(* Logix 5000 project; controller POA Emulate 5570 rev 30.12; software revision 30.00 *)

TASK MainTask (periodic, rate 10000 ms, priority 1, watchdog 10000 ms) : MainProgram

MODULES
   Local : Emulate 5570 (ICP 2, rev 30.12)
END_MODULES

VAR_GLOBAL   (* controller tags *)
   _SEC_P : BOOL;
   done : DINT;
   R_TRIG : FBD_ONESHOT;
   temp_var : DINT;
   test_array : DINT[20] := ([0] := 1, [1] := 2, [2] := 3, [3] := 4, [4] := 5, [5] := 6, [6] := 7, [7] := 8, [8] := 9, [9] := 10, [10] := 11, [11] := 12, [12] := 13, [13] := 14, [14] := 15, [15] := 16, [16] := 17, [17] := 18, [18] := 19, [19] := 20);
   TON : FBD_TIMER;
END_VAR

PROGRAM MainProgram   (* main routine MainRoutine *)
VAR
   Chaskey_128_i : DINT;
   Chaskey_a : DINT; {access None}
   Chaskey_BNum : DINT; {access None}
   Chaskey_i : DINT; {access None}
   Chaskey_IndexDiv : DINT;
   Chaskey_IndexMod : DINT;
   Chaskey_input_pi : DINT[4]; {access None}
   Chaskey_j : DINT; {access None}
   Chaskey_key : DINT[4]; {access None}
   Chaskey_L : DINT[4]; {access None}
   Chaskey_LastBlk : DINT[4];
   Chaskey_lb : DINT[16];
   Chaskey_Message : DINT[256]; {access None}
   Chaskey_mlen : DINT;
   Chaskey_MsgBitLen : DINT;
   Chaskey_MsgBlk : DINT[16];
   Chaskey_MsgBlkLen : DINT;
   Chaskey_per_i : DINT; {access None}
   Chaskey_round : DINT;
   Chaskey_shift_input : DINT; {access None}
   Chaskey_shift_result : DINT; {access None}
   Chaskey_subkey1_i : DINT; {access None}
   Chaskey_subkey2_i : DINT; {access None}
   Chaskey_subkey_1 : DINT[8];
   Chaskey_subkey_2 : DINT[8]; {access None}
   Chaskey_tag : DINT[4]; {access None}
   Chaskey_Temp : DINT; {access None}
   Chaskey_z : DINT;
   Date_time : DINT[7]; {access None}
        [0]   // Year
        [1]   // Month
        [2]   // Day
        [3]   // Hour
        [4]   // Minute
        [5]   // Second
        [6]   // Microsecond
   OWF_Add_c : DINT;
   OWF_i : DINT;
   OWF_Input : DINT[17];
   OWF_InputLen : DINT;
   OWF_InputMaxInd : DINT;
   OWF_Result : DINT[17];
   POA_Chain_NM : DINT; {access None}
   POA_CK_RefillNM : DINT; {access None}
   POA_CKP : DINT[17]; {access None}
   POA_CKP_Ctx : DINT[9,16]; {access None}
   POA_CKP_Indx : DINT[9]; {access None}
   POA_i : DINT;
   POA_Ins_NM : DINT; {access None}
   POA_is_Bootstrap : BOOL; {access None}
   POA_j : DINT;
   POA_k : DINT; {access None}
   POA_lr : DINT;
   POA_m : DINT;
   POA_Microsecond1 : DINT; {access None}
   POA_Microsecond2 : DINT; {access None}
   POA_MicrosecondABS : DINT;
   POA_OTS : SINT[256,256];
   POA_Pf : DINT[17]; {access None}
   POA_Pf_Indx : DINT; {access None}
   PoA_Pf_Interval : DINT;
   POA_Qu_head : DINT; {access None}
   POA_Qu_tail : DINT; {access None}
   POA_SC_DeltaS : DINT;
   POA_SC_Interval : DINT;
   POA_Second1 : DINT; {access None}
   POA_Second2 : DINT; {access None}
   POA_SecondABS : DINT;
   POA_SIG_i : DINT;
   POA_tag : DINT[4]; {access None}
   POA_Vrf_Points : DINT[260,17];
   PRG_Counter : DINT[2];
   PRG_i : DINT;
   PRG_j : DINT;
   PRG_Res_Len : DINT;
   PRG_Result : DINT[128];
   SCAN_CYCLE_TIME : DINT; {access None}
   UOWHF_Add_c : DINT;
   UOWHF_i : DINT;
   UOWHF_InputLen : DINT;
   UOWHF_InputMaxInd : DINT := 7;
   UOWHF_Msg : DINT[17];
   UOWHF_OutputMaxInd : DINT;
   UOWHF_Result : DINT[17];
   UOWHF_Vary_BlkNum : DINT;
   UOWHF_Vary_i : DINT := 256;
   UOWHF_Vary_j : DINT;
   UOWHF_Vary_Message : DINT[3000] := ([0] := 1, [1] := 1, [2] := 1, [3] := 1, [4] := 1, [5] := 1, [6] := 1, [7] := 1, [8] := 1, [9] := 1, [10] := 1, [11] := 1, [12] := 1, [13] := 1, [14] := 1, [15] := 1, [16] := 1, [17] := 1, [18] := 1, [19] := 1, [20] := 1, [21] := 1, [22] := 1, [23] := 1, [24] := 1, [25] := 1, [26] := 1, [27] := 1, [28] := 1, [29] := 1, [30] := 1, [31] := 1, [32] := 1, [33] := 1, [34] := 1, [35] := 1, [36] := 1, [37] := 1, [38] := 1, [39] := 1, [40] := 1, [41] := 1, [42] := 1, [43] := 1, [44] := 1, [45] := 1, [46] := 1, [47] := 1, [48] := 1, [49] := 1, [50] := 1, [51] := 1, [52] := 1, [53] := 1, [54] := 1, [55] := 1, [56] := 1, [57] := 1, [58] := 1, [59] := 1,
        [60] := 1, [61] := 1, [62] := 1, [63] := 1, [64] := 1, [65] := 1, [66] := 1, [67] := 1, [68] := 1, [69] := 1, [70] := 1, [71] := 1, [72] := 1, [73] := 1, [74] := 1, [75] := 1, [76] := 1, [77] := 1, [78] := 1, [79] := 1, [80] := 1, [81] := 1, [82] := 1, [83] := 1, [84] := 1, [85] := 1, [86] := 1, [87] := 1, [88] := 1, [89] := 1, [90] := 1, [91] := 1, [92] := 1, [93] := 1, [94] := 1, [95] := 1, [96] := 1, [97] := 1, [98] := 1, [99] := 1, [100] := 1, [101] := 1, [102] := 1, [103] := 1, [104] := 1, [105] := 1, [106] := 1, [107] := 1, [108] := 1, [109] := 1, [110] := 1, [111] := 1, [112] := 1, [113] := 1, [114] := 1, [115] := 1, [116] := 1, [117] := 1, [118] := 1, [119] := 1,
        [120] := 1, [121] := 1, [122] := 1, [123] := 1, [124] := 1, [125] := 1, [126] := 1, [127] := 1, [128] := 1, [129] := 1, [130] := 1, [131] := 1, [132] := 1, [133] := 1, [134] := 1, [135] := 1, [136] := 1, [137] := 1, [138] := 1, [139] := 1, [140] := 1, [141] := 1, [142] := 1, [143] := 1, [144] := 1, [145] := 1, [146] := 1, [147] := 1, [148] := 1, [149] := 1, [150] := 1, [151] := 1, [152] := 1, [153] := 1, [154] := 1, [155] := 1, [156] := 1, [157] := 1, [158] := 1, [159] := 1, [160] := 1, [161] := 1, [162] := 1, [163] := 1, [164] := 1, [165] := 1, [166] := 1, [167] := 1, [168] := 1, [169] := 1, [170] := 1, [171] := 1, [172] := 1, [173] := 1, [174] := 1, [175] := 1, [176] := 1, [177] := 1, [178] := 1, [179] := 1,
        [180] := 1, [181] := 1, [182] := 1, [183] := 1, [184] := 1, [185] := 1, [186] := 1, [187] := 1, [188] := 1, [189] := 1, [190] := 1, [191] := 1, [192] := 1, [193] := 1, [194] := 1, [195] := 1, [196] := 1, [197] := 1, [198] := 1, [199] := 1, [200] := 1, [201] := 1, [202] := 1, [203] := 1, [204] := 1, [205] := 1, [206] := 1, [207] := 1, [208] := 1, [209] := 1, [210] := 1, [211] := 1, [212] := 1, [213] := 1, [214] := 1, [215] := 1, [216] := 1, [217] := 1, [218] := 1, [219] := 1, [220] := 1, [221] := 1, [222] := 1, [223] := 1, [224] := 1, [225] := 1, [226] := 1, [227] := 1, [228] := 1, [229] := 1, [230] := 1, [231] := 1, [232] := 1, [233] := 1, [234] := 1, [235] := 1, [236] := 1, [237] := 1, [238] := 1, [239] := 1,
        [240] := 1, [241] := 1, [242] := 1, [243] := 1, [244] := 1, [245] := 1, [246] := 1, [247] := 1, [248] := 1, [249] := 1, [250] := 1, [251] := 1, [252] := 1, [253] := 1, [254] := 1, [255] := 1);
   UOWHF_Vary_MsgLen : DINT := 255;
   UOWHF_Vary_OutputMaxInd : DINT := 4;
   UOWHF_Vary_z : DINT;
   UOWHF_VaryLen : DINT;
   UOWHF_Ver : DINT;
END_VAR

ROUTINE Application   (* structured text *)
   //Description: initialize the variables.
   
   if S:FS then  (* this is the first, normal scan of the routines in the current program, initialize the program.*)
   
   
   
   
   
   end_if;
   
   
   
   
   
END_ROUTINE

ROUTINE CHASKEY_128   (* structured text *)
   JSR(CHASKEY_Init);
   
   Chaskey_BNum:= Chaskey_MsgBitLen/128;
   
   if Chaskey_MsgBitLen mod 128 <>0 then
   	Chaskey_BNum:= Chaskey_BNum+1;
   end_if;
   
   
   for Chaskey_i:=0 to Chaskey_mlen by 1 do
   	Chaskey_MsgBlkLen:=Chaskey_mlen/4;
   	Chaskey_z:=Chaskey_i mod 4;
   	for Chaskey_j:=0 to 7 by 1 do
   		Chaskey_MsgBlk[Chaskey_MsgBlkLen].[Chaskey_z*8+Chaskey_j]:=Chaskey_Message[Chaskey_i].[Chaskey_j];
   	end_for;
   end_for;
   
   Chaskey_input_pi[3] := Chaskey_key[3];
   Chaskey_input_pi[2] := Chaskey_key[2] ;
   Chaskey_input_pi[1] := Chaskey_key[1] ;
   Chaskey_input_pi[0] := Chaskey_key[0] ;
   
   Chaskey_i:=0;
   if Chaskey_mlen<>0 then
   	while Chaskey_i < Chaskey_BNum-1 do
   		Chaskey_128_i:=Chaskey_i*4;
   		Chaskey_input_pi[3] := Chaskey_input_pi[3] XOR Chaskey_MsgBlk[Chaskey_128_i+3];
   		Chaskey_input_pi[2] := Chaskey_input_pi[2] XOR Chaskey_MsgBlk[Chaskey_128_i+2];
   		Chaskey_input_pi[1] := Chaskey_input_pi[1] XOR Chaskey_MsgBlk[Chaskey_128_i+1];
   		Chaskey_input_pi[0] := Chaskey_input_pi[0] XOR Chaskey_MsgBlk[Chaskey_128_i+0];
   		JSR(CHASKEY_Permutation);
   
   		if Chaskey_i>=Chaskey_BNum-2 then
   			Exit;
   		end_if;
   
   		Chaskey_i:=Chaskey_i +1;
   	end_while;
   end_if;
   
   
   if (Chaskey_mlen<>0) AND ((Chaskey_mlen & 15)=0) then
   	Chaskey_L[3] := Chaskey_subkey_1[3];
   	Chaskey_L[2] := Chaskey_subkey_1[2] ;
   	Chaskey_L[1] := Chaskey_subkey_1[1] ;
   	Chaskey_L[0] := Chaskey_subkey_1[0] ;
   	Chaskey_LastBlk[0]:=Chaskey_MsgBlk[0];
   	Chaskey_LastBlk[1]:=Chaskey_MsgBlk[1];
   	Chaskey_LastBlk[2]:=Chaskey_MsgBlk[2];
   	Chaskey_LastBlk[3]:=Chaskey_MsgBlk[3];
   else
   	Chaskey_L[3] := Chaskey_subkey_2[3];
   	Chaskey_L[2] := Chaskey_subkey_2[2] ;
   	Chaskey_L[1] := Chaskey_subkey_2[1] ;
   	Chaskey_L[0] := Chaskey_subkey_2[0] ;
   
   
   	Chaskey_IndexMod:= Chaskey_mlen mod 16;
   	Chaskey_IndexDiv:= (Chaskey_mlen/16)*16;
   	for Chaskey_j:=0 to Chaskey_IndexMod-1 by 1 do
   		Chaskey_lb[Chaskey_j]:=Chaskey_Message[Chaskey_IndexDiv+Chaskey_j];
   	end_for;
   	Chaskey_lb[Chaskey_IndexMod]:=1;
   	for Chaskey_j:=Chaskey_IndexMod+1 to 15 by 1 do
   		Chaskey_lb[Chaskey_j]:=0;
   	end_for;
   
   	//lastblock = (uint32_t*) lb;
   	Chaskey_LastBlk[0].0:=Chaskey_lb[0].0;
   	Chaskey_LastBlk[0].1:=Chaskey_lb[0].1;
   	Chaskey_LastBlk[0].2:=Chaskey_lb[0].2;
   	Chaskey_LastBlk[0].3:=Chaskey_lb[0].3;
   	Chaskey_LastBlk[0].4:=Chaskey_lb[0].4;
   	Chaskey_LastBlk[0].5:=Chaskey_lb[0].5;
   	Chaskey_LastBlk[0].6:=Chaskey_lb[0].6;
   	Chaskey_LastBlk[0].7:=Chaskey_lb[0].7;
   	Chaskey_LastBlk[0].8:=Chaskey_lb[1].0;
   	Chaskey_LastBlk[0].9:=Chaskey_lb[1].1;
   	Chaskey_LastBlk[0].10:=Chaskey_lb[1].2;
   	Chaskey_LastBlk[0].11:=Chaskey_lb[1].3;
   	Chaskey_LastBlk[0].12:=Chaskey_lb[1].4;
   	Chaskey_LastBlk[0].13:=Chaskey_lb[1].5;
   	Chaskey_LastBlk[0].14:=Chaskey_lb[1].6;
   	Chaskey_LastBlk[0].15:=Chaskey_lb[1].7;
   	Chaskey_LastBlk[0].16:=Chaskey_lb[2].0;
   	Chaskey_LastBlk[0].17:=Chaskey_lb[2].1;
   	Chaskey_LastBlk[0].18:=Chaskey_lb[2].2;
   	Chaskey_LastBlk[0].19:=Chaskey_lb[2].3;
   	Chaskey_LastBlk[0].20:=Chaskey_lb[2].4;
   	Chaskey_LastBlk[0].21:=Chaskey_lb[2].5;
   	Chaskey_LastBlk[0].22:=Chaskey_lb[2].6;
   	Chaskey_LastBlk[0].23:=Chaskey_lb[2].7;
   	Chaskey_LastBlk[0].24:=Chaskey_lb[3].0;
   	Chaskey_LastBlk[0].25:=Chaskey_lb[3].1;
   	Chaskey_LastBlk[0].26:=Chaskey_lb[3].2;
   	Chaskey_LastBlk[0].27:=Chaskey_lb[3].3;
   	Chaskey_LastBlk[0].28:=Chaskey_lb[3].4;
   	Chaskey_LastBlk[0].29:=Chaskey_lb[3].5;
   	Chaskey_LastBlk[0].30:=Chaskey_lb[3].6;
   	Chaskey_LastBlk[0].31:=Chaskey_lb[3].7;
   
   	Chaskey_LastBlk[1].0:=Chaskey_lb[4].0;
   	Chaskey_LastBlk[1].1:=Chaskey_lb[4].1;
   	Chaskey_LastBlk[1].2:=Chaskey_lb[4].2;
   	Chaskey_LastBlk[1].3:=Chaskey_lb[4].3;
   	Chaskey_LastBlk[1].4:=Chaskey_lb[4].4;
   	Chaskey_LastBlk[1].5:=Chaskey_lb[4].5;
   	Chaskey_LastBlk[1].6:=Chaskey_lb[4].6;
   	Chaskey_LastBlk[1].7:=Chaskey_lb[4].7;
   	Chaskey_LastBlk[1].8:=Chaskey_lb[5].0;
   	Chaskey_LastBlk[1].9:=Chaskey_lb[5].1;
   	Chaskey_LastBlk[1].10:=Chaskey_lb[5].2;
   	Chaskey_LastBlk[1].11:=Chaskey_lb[5].3;
   	Chaskey_LastBlk[1].12:=Chaskey_lb[5].4;
   	Chaskey_LastBlk[1].13:=Chaskey_lb[5].5;
   	Chaskey_LastBlk[1].14:=Chaskey_lb[5].6;
   	Chaskey_LastBlk[1].15:=Chaskey_lb[5].7;
   	Chaskey_LastBlk[1].16:=Chaskey_lb[6].0;
   	Chaskey_LastBlk[1].17:=Chaskey_lb[6].1;
   	Chaskey_LastBlk[1].18:=Chaskey_lb[6].2;
   	Chaskey_LastBlk[1].19:=Chaskey_lb[6].3;
   	Chaskey_LastBlk[1].20:=Chaskey_lb[6].4;
   	Chaskey_LastBlk[1].21:=Chaskey_lb[6].5;
   	Chaskey_LastBlk[1].22:=Chaskey_lb[6].6;
   	Chaskey_LastBlk[1].23:=Chaskey_lb[6].7;
   	Chaskey_LastBlk[1].24:=Chaskey_lb[7].0;
   	Chaskey_LastBlk[1].25:=Chaskey_lb[7].1;
   	Chaskey_LastBlk[1].26:=Chaskey_lb[7].2;
   	Chaskey_LastBlk[1].27:=Chaskey_lb[7].3;
   	Chaskey_LastBlk[1].28:=Chaskey_lb[7].4;
   	Chaskey_LastBlk[1].29:=Chaskey_lb[7].5;
   	Chaskey_LastBlk[1].30:=Chaskey_lb[7].6;
   	Chaskey_LastBlk[1].31:=Chaskey_lb[7].7;
   
   	Chaskey_LastBlk[2].0:=Chaskey_lb[8].0;
   	Chaskey_LastBlk[2].1:=Chaskey_lb[8].1;
   	Chaskey_LastBlk[2].2:=Chaskey_lb[8].2;
   	Chaskey_LastBlk[2].3:=Chaskey_lb[8].3;
   	Chaskey_LastBlk[2].4:=Chaskey_lb[8].4;
   	Chaskey_LastBlk[2].5:=Chaskey_lb[8].5;
   	Chaskey_LastBlk[2].6:=Chaskey_lb[8].6;
   	Chaskey_LastBlk[2].7:=Chaskey_lb[8].7;
   	Chaskey_LastBlk[2].8:=Chaskey_lb[9].0;
   	Chaskey_LastBlk[2].9:=Chaskey_lb[9].1;
   	Chaskey_LastBlk[2].10:=Chaskey_lb[9].2;
   	Chaskey_LastBlk[2].11:=Chaskey_lb[9].3;
   	Chaskey_LastBlk[2].12:=Chaskey_lb[9].4;
   	Chaskey_LastBlk[2].13:=Chaskey_lb[9].5;
   	Chaskey_LastBlk[2].14:=Chaskey_lb[9].6;
   	Chaskey_LastBlk[2].15:=Chaskey_lb[9].7;
   	Chaskey_LastBlk[2].16:=Chaskey_lb[10].0;
   	Chaskey_LastBlk[2].17:=Chaskey_lb[10].1;
   	Chaskey_LastBlk[2].18:=Chaskey_lb[10].2;
   	Chaskey_LastBlk[2].19:=Chaskey_lb[10].3;
   	Chaskey_LastBlk[2].20:=Chaskey_lb[10].4;
   	Chaskey_LastBlk[2].21:=Chaskey_lb[10].5;
   	Chaskey_LastBlk[2].22:=Chaskey_lb[10].6;
   	Chaskey_LastBlk[2].23:=Chaskey_lb[10].7;
   	Chaskey_LastBlk[2].24:=Chaskey_lb[11].0;
   	Chaskey_LastBlk[2].25:=Chaskey_lb[11].1;
   	Chaskey_LastBlk[2].26:=Chaskey_lb[11].2;
   	Chaskey_LastBlk[2].27:=Chaskey_lb[11].3;
   	Chaskey_LastBlk[2].28:=Chaskey_lb[11].4;
   	Chaskey_LastBlk[2].29:=Chaskey_lb[11].5;
   	Chaskey_LastBlk[2].30:=Chaskey_lb[11].6;
   	Chaskey_LastBlk[2].31:=Chaskey_lb[11].7;
   
   	Chaskey_LastBlk[3].0:=Chaskey_lb[12].0;
   	Chaskey_LastBlk[3].1:=Chaskey_lb[12].1;
   	Chaskey_LastBlk[3].2:=Chaskey_lb[12].2;
   	Chaskey_LastBlk[3].3:=Chaskey_lb[12].3;
   	Chaskey_LastBlk[3].4:=Chaskey_lb[12].4;
   	Chaskey_LastBlk[3].5:=Chaskey_lb[12].5;
   	Chaskey_LastBlk[3].6:=Chaskey_lb[12].6;
   	Chaskey_LastBlk[3].7:=Chaskey_lb[12].7;
   	Chaskey_LastBlk[3].8:=Chaskey_lb[13].0;
   	Chaskey_LastBlk[3].9:=Chaskey_lb[13].1;
   	Chaskey_LastBlk[3].10:=Chaskey_lb[13].2;
   	Chaskey_LastBlk[3].11:=Chaskey_lb[13].3;
   	Chaskey_LastBlk[3].12:=Chaskey_lb[13].4;
   	Chaskey_LastBlk[3].13:=Chaskey_lb[13].5;
   	Chaskey_LastBlk[3].14:=Chaskey_lb[13].6;
   	Chaskey_LastBlk[3].15:=Chaskey_lb[13].7;
   	Chaskey_LastBlk[3].16:=Chaskey_lb[14].0;
   	Chaskey_LastBlk[3].17:=Chaskey_lb[14].1;
   	Chaskey_LastBlk[3].18:=Chaskey_lb[14].2;
   	Chaskey_LastBlk[3].19:=Chaskey_lb[14].3;
   	Chaskey_LastBlk[3].20:=Chaskey_lb[14].4;
   	Chaskey_LastBlk[3].21:=Chaskey_lb[14].5;
   	Chaskey_LastBlk[3].22:=Chaskey_lb[14].6;
   	Chaskey_LastBlk[3].23:=Chaskey_lb[14].7;
   	Chaskey_LastBlk[3].24:=Chaskey_lb[15].0;
   	Chaskey_LastBlk[3].25:=Chaskey_lb[15].1;
   	Chaskey_LastBlk[3].26:=Chaskey_lb[15].2;
   	Chaskey_LastBlk[3].27:=Chaskey_lb[15].3;
   	Chaskey_LastBlk[3].28:=Chaskey_lb[15].4;
   	Chaskey_LastBlk[3].29:=Chaskey_lb[15].5;
   	Chaskey_LastBlk[3].30:=Chaskey_lb[15].6;
   	Chaskey_LastBlk[3].31:=Chaskey_lb[15].7;
   end_if;
   
   
   Chaskey_input_pi[3] := Chaskey_input_pi[3] XOR Chaskey_LastBlk[3] ;
   Chaskey_input_pi[2] := Chaskey_input_pi[2] XOR Chaskey_LastBlk[2] ;
   Chaskey_input_pi[1] := Chaskey_input_pi[1] XOR Chaskey_LastBlk[1] ;
   Chaskey_input_pi[0] := Chaskey_input_pi[0] XOR Chaskey_LastBlk[0] ;
   
   Chaskey_input_pi[3] := Chaskey_input_pi[3] XOR Chaskey_L[3] ;
   Chaskey_input_pi[2] := Chaskey_input_pi[2] XOR Chaskey_L[2] ;
   Chaskey_input_pi[1] := Chaskey_input_pi[1] XOR Chaskey_L[1] ;
   Chaskey_input_pi[0] := Chaskey_input_pi[0] XOR Chaskey_L[0] ;
   
   JSR(CHASKEY_Permutation);
   
   Chaskey_input_pi[3] := Chaskey_input_pi[3] XOR Chaskey_L[3] ;
   Chaskey_input_pi[2] := Chaskey_input_pi[2] XOR Chaskey_L[2] ;
   Chaskey_input_pi[1] := Chaskey_input_pi[1] XOR Chaskey_L[1] ;
   Chaskey_input_pi[0] := Chaskey_input_pi[0] XOR Chaskey_L[0] ;
   
   //////////////////////////////////////////////
   
   Chaskey_tag[3] := Chaskey_input_pi[3];
   Chaskey_tag[2] := Chaskey_input_pi[2];
   Chaskey_tag[1] := Chaskey_input_pi[1];
   Chaskey_tag[0] := Chaskey_input_pi[0];
   
   JSR(CHASKEY_ClearKey);
   
END_ROUTINE

ROUTINE CHASKEY_ClearKey   (* structured text *)
   
   Chaskey_key[0]:= 0;
   Chaskey_key[1]:= 0;
   Chaskey_key[2]:= 0;
   Chaskey_key[3]:= 0;
   
   Chaskey_subkey_1[0]:= 0;
   Chaskey_subkey_1[1]:= 0;
   Chaskey_subkey_1[2]:= 0;
   Chaskey_subkey_1[3]:= 0;
   
   Chaskey_subkey_2[0]:= 0;
   Chaskey_subkey_2[1]:= 0;
   Chaskey_subkey_2[2]:= 0;
   Chaskey_subkey_2[3]:= 0;
   
END_ROUTINE

ROUTINE CHASKEY_Init   (* structured text *)
    //key[3].31 is the MSB of the key, while key[0].0 is the LSB of the key
   (*Chaskey_key[0]:=0;
   Chaskey_key[1]:=17;
   Chaskey_key[2]:=34;
   Chaskey_key[3]:=51;*)
   
   Chaskey_key[0]:=857870592;
   Chaskey_key[1]:=2003195204;
   Chaskey_key[2]:=-1146447480;
   Chaskey_key[3]:=-1122868;
   
   Chaskey_tag[0] := 0;
   Chaskey_tag[1] := 0;
   Chaskey_tag[2] := 0;
   Chaskey_tag[3] := 0;
   
   //Initialize subkey_1[] and subkey_2[]
   Chaskey_subkey_1[0] := 1715741319;
   Chaskey_subkey_1[1] := -288576888;
   Chaskey_subkey_1[2] := 2002070336;
   Chaskey_subkey_1[3] := -2245735;
   
   Chaskey_subkey_2[0] := -863484535;
   Chaskey_subkey_2[1] := -577153776;
   Chaskey_subkey_2[2] := -290822623;
   Chaskey_subkey_2[3] := -4491470;
   
   
   
END_ROUTINE

ROUTINE CHASKEY_Permutation   (* structured text *)
   
   for Chaskey_per_i:=0 to Chaskey_round by 1 do
   
   
   	Chaskey_input_pi[0]:= Chaskey_input_pi[0] + Chaskey_input_pi[1];
   
   	Chaskey_a:=Chaskey_input_pi[1];  //v1 <<< 5
   	Chaskey_Temp:=0;
   	//left shift Chaskey_b=5 bits
   	Chaskey_Temp.5:=Chaskey_a.0;
   	Chaskey_Temp.6:=Chaskey_a.1;
   	Chaskey_Temp.7:=Chaskey_a.2;
   	Chaskey_Temp.8:=Chaskey_a.3;
   	Chaskey_Temp.9:=Chaskey_a.4;
   	Chaskey_Temp.10:=Chaskey_a.5;
   	Chaskey_Temp.11:=Chaskey_a.6;
   	Chaskey_Temp.12:=Chaskey_a.7;
   	Chaskey_Temp.13:=Chaskey_a.8;
   	Chaskey_Temp.14:=Chaskey_a.9;
   	Chaskey_Temp.15:=Chaskey_a.10;
   	Chaskey_Temp.16:=Chaskey_a.11;
   	Chaskey_Temp.17:=Chaskey_a.12;
   	Chaskey_Temp.18:=Chaskey_a.13;
   	Chaskey_Temp.19:=Chaskey_a.14;
   	Chaskey_Temp.20:=Chaskey_a.15;
   	Chaskey_Temp.21:=Chaskey_a.16;
   	Chaskey_Temp.22:=Chaskey_a.17;
   	Chaskey_Temp.23:=Chaskey_a.18;
   	Chaskey_Temp.24:=Chaskey_a.19;
   	Chaskey_Temp.25:=Chaskey_a.20;
   	Chaskey_Temp.26:=Chaskey_a.21;
   	Chaskey_Temp.27:=Chaskey_a.22;
   	Chaskey_Temp.28:=Chaskey_a.23;
   	Chaskey_Temp.29:=Chaskey_a.24;
   	Chaskey_Temp.30:=Chaskey_a.25;
   	Chaskey_Temp.31:=Chaskey_a.26;
   	Chaskey_Temp.0:=Chaskey_a.27;
   	Chaskey_Temp.1:=Chaskey_a.28;
   	Chaskey_Temp.2:=Chaskey_a.29;
   	Chaskey_Temp.3:=Chaskey_a.30;
   	Chaskey_Temp.4:=Chaskey_a.31;
   	Chaskey_input_pi[1]:=Chaskey_Temp;
   
   	Chaskey_input_pi[1]:=Chaskey_input_pi[1] XOR Chaskey_input_pi[0];
   
   
   	Chaskey_a:=Chaskey_input_pi[0];  // <<< 16
   	Chaskey_Temp:=0;
   	//left shift Chaskey_b=16 bits
   	Chaskey_Temp.16:=Chaskey_a.0;
   	Chaskey_Temp.17:=Chaskey_a.1;
   	Chaskey_Temp.18:=Chaskey_a.2;
   	Chaskey_Temp.19:=Chaskey_a.3;
   	Chaskey_Temp.20:=Chaskey_a.4;
   	Chaskey_Temp.21:=Chaskey_a.5;
   	Chaskey_Temp.22:=Chaskey_a.6;
   	Chaskey_Temp.23:=Chaskey_a.7;
   	Chaskey_Temp.24:=Chaskey_a.8;
   	Chaskey_Temp.25:=Chaskey_a.9;
   	Chaskey_Temp.26:=Chaskey_a.10;
   	Chaskey_Temp.27:=Chaskey_a.11;
   	Chaskey_Temp.28:=Chaskey_a.12;
   	Chaskey_Temp.29:=Chaskey_a.13;
   	Chaskey_Temp.30:=Chaskey_a.14;
   	Chaskey_Temp.31:=Chaskey_a.15;
   	Chaskey_Temp.0:=Chaskey_a.16;
   	Chaskey_Temp.1:=Chaskey_a.17;
   	Chaskey_Temp.2:=Chaskey_a.18;
   	Chaskey_Temp.3:=Chaskey_a.19;
   	Chaskey_Temp.4:=Chaskey_a.20;
   	Chaskey_Temp.5:=Chaskey_a.21;
   	Chaskey_Temp.6:=Chaskey_a.22;
   	Chaskey_Temp.7:=Chaskey_a.23;
   	Chaskey_Temp.8:=Chaskey_a.24;
   	Chaskey_Temp.9:=Chaskey_a.25;
   	Chaskey_Temp.10:=Chaskey_a.26;
   	Chaskey_Temp.11:=Chaskey_a.27;
   	Chaskey_Temp.12:=Chaskey_a.28;
   	Chaskey_Temp.13:=Chaskey_a.29;
   	Chaskey_Temp.14:=Chaskey_a.30;
   	Chaskey_Temp.15:=Chaskey_a.31;
   	Chaskey_input_pi[0]:=Chaskey_Temp;
   
   
       Chaskey_input_pi[2]:= Chaskey_input_pi[2] + Chaskey_input_pi[3];
   
   
   	Chaskey_a:=Chaskey_input_pi[3];  // <<< 8
   	Chaskey_Temp:=0;
   	//left shift Chaskey_b=8 bits
   	Chaskey_Temp.8:=Chaskey_a.0;
   	Chaskey_Temp.9:=Chaskey_a.1;
   	Chaskey_Temp.10:=Chaskey_a.2;
   	Chaskey_Temp.11:=Chaskey_a.3;
   	Chaskey_Temp.12:=Chaskey_a.4;
   	Chaskey_Temp.13:=Chaskey_a.5;
   	Chaskey_Temp.14:=Chaskey_a.6;
   	Chaskey_Temp.15:=Chaskey_a.7;
   	Chaskey_Temp.16:=Chaskey_a.8;
   	Chaskey_Temp.17:=Chaskey_a.9;
   	Chaskey_Temp.18:=Chaskey_a.10;
   	Chaskey_Temp.19:=Chaskey_a.11;
   	Chaskey_Temp.20:=Chaskey_a.12;
   	Chaskey_Temp.21:=Chaskey_a.13;
   	Chaskey_Temp.22:=Chaskey_a.14;
   	Chaskey_Temp.23:=Chaskey_a.15;
   	Chaskey_Temp.24:=Chaskey_a.16;
   	Chaskey_Temp.25:=Chaskey_a.17;
   	Chaskey_Temp.26:=Chaskey_a.18;
   	Chaskey_Temp.27:=Chaskey_a.19;
   	Chaskey_Temp.28:=Chaskey_a.20;
   	Chaskey_Temp.29:=Chaskey_a.21;
   	Chaskey_Temp.30:=Chaskey_a.22;
   	Chaskey_Temp.31:=Chaskey_a.23;
   	Chaskey_Temp.0:=Chaskey_a.24;
   	Chaskey_Temp.1:=Chaskey_a.25;
   	Chaskey_Temp.2:=Chaskey_a.26;
   	Chaskey_Temp.3:=Chaskey_a.27;
   	Chaskey_Temp.4:=Chaskey_a.28;
   	Chaskey_Temp.5:=Chaskey_a.29;
   	Chaskey_Temp.6:=Chaskey_a.30;
   	Chaskey_Temp.7:=Chaskey_a.31;
   	Chaskey_input_pi[3]:=Chaskey_Temp;
   
   	Chaskey_input_pi[3]:=Chaskey_input_pi[3] XOR Chaskey_input_pi[2];
   
   
   
   	Chaskey_input_pi[0]:= Chaskey_input_pi[0] + Chaskey_input_pi[3];
   
   	Chaskey_a:=Chaskey_input_pi[3];  //<<< 13
   	Chaskey_Temp:=0;
   	//left shift Chaskey_b=13 bits
   	Chaskey_Temp.13:=Chaskey_a.0;
   	Chaskey_Temp.14:=Chaskey_a.1;
   	Chaskey_Temp.15:=Chaskey_a.2;
   	Chaskey_Temp.16:=Chaskey_a.3;
   	Chaskey_Temp.17:=Chaskey_a.4;
   	Chaskey_Temp.18:=Chaskey_a.5;
   	Chaskey_Temp.19:=Chaskey_a.6;
   	Chaskey_Temp.20:=Chaskey_a.7;
   	Chaskey_Temp.21:=Chaskey_a.8;
   	Chaskey_Temp.22:=Chaskey_a.9;
   	Chaskey_Temp.23:=Chaskey_a.10;
   	Chaskey_Temp.24:=Chaskey_a.11;
   	Chaskey_Temp.25:=Chaskey_a.12;
   	Chaskey_Temp.26:=Chaskey_a.13;
   	Chaskey_Temp.27:=Chaskey_a.14;
   	Chaskey_Temp.28:=Chaskey_a.15;
   	Chaskey_Temp.29:=Chaskey_a.16;
   	Chaskey_Temp.30:=Chaskey_a.17;
   	Chaskey_Temp.31:=Chaskey_a.18;
   	Chaskey_Temp.0:=Chaskey_a.19;
   	Chaskey_Temp.1:=Chaskey_a.20;
   	Chaskey_Temp.2:=Chaskey_a.21;
   	Chaskey_Temp.3:=Chaskey_a.22;
   	Chaskey_Temp.4:=Chaskey_a.23;
   	Chaskey_Temp.5:=Chaskey_a.24;
   	Chaskey_Temp.6:=Chaskey_a.25;
   	Chaskey_Temp.7:=Chaskey_a.26;
   	Chaskey_Temp.8:=Chaskey_a.27;
   	Chaskey_Temp.9:=Chaskey_a.28;
   	Chaskey_Temp.10:=Chaskey_a.29;
   	Chaskey_Temp.11:=Chaskey_a.30;
   	Chaskey_Temp.12:=Chaskey_a.31;
   	Chaskey_input_pi[3]:=Chaskey_Temp;
   
   	Chaskey_input_pi[3]:=Chaskey_input_pi[3] XOR Chaskey_input_pi[0];
   
   
   	Chaskey_input_pi[2]:=  Chaskey_input_pi[2] + Chaskey_input_pi[1];
   
   	Chaskey_a:=Chaskey_input_pi[1]; //<<< 7
   	Chaskey_Temp:=0;
   	//left shift Chaskey_b=7 bits
   	Chaskey_Temp.7:=Chaskey_a.0;
   	Chaskey_Temp.8:=Chaskey_a.1;
   	Chaskey_Temp.9:=Chaskey_a.2;
   	Chaskey_Temp.10:=Chaskey_a.3;
   	Chaskey_Temp.11:=Chaskey_a.4;
   	Chaskey_Temp.12:=Chaskey_a.5;
   	Chaskey_Temp.13:=Chaskey_a.6;
   	Chaskey_Temp.14:=Chaskey_a.7;
   	Chaskey_Temp.15:=Chaskey_a.8;
   	Chaskey_Temp.16:=Chaskey_a.9;
   	Chaskey_Temp.17:=Chaskey_a.10;
   	Chaskey_Temp.18:=Chaskey_a.11;
   	Chaskey_Temp.19:=Chaskey_a.12;
   	Chaskey_Temp.20:=Chaskey_a.13;
   	Chaskey_Temp.21:=Chaskey_a.14;
   	Chaskey_Temp.22:=Chaskey_a.15;
   	Chaskey_Temp.23:=Chaskey_a.16;
   	Chaskey_Temp.24:=Chaskey_a.17;
   	Chaskey_Temp.25:=Chaskey_a.18;
   	Chaskey_Temp.26:=Chaskey_a.19;
   	Chaskey_Temp.27:=Chaskey_a.20;
   	Chaskey_Temp.28:=Chaskey_a.21;
   	Chaskey_Temp.29:=Chaskey_a.22;
   	Chaskey_Temp.30:=Chaskey_a.23;
   	Chaskey_Temp.31:=Chaskey_a.24;
   	Chaskey_Temp.0:=Chaskey_a.25;
   	Chaskey_Temp.1:=Chaskey_a.26;
   	Chaskey_Temp.2:=Chaskey_a.27;
   	Chaskey_Temp.3:=Chaskey_a.28;
   	Chaskey_Temp.4:=Chaskey_a.29;
   	Chaskey_Temp.5:=Chaskey_a.30;
   	Chaskey_Temp.6:=Chaskey_a.31;
   	Chaskey_input_pi[1]:=Chaskey_Temp;
   
   	Chaskey_input_pi[1]:=Chaskey_input_pi[1] XOR Chaskey_input_pi[2];
   
   
   	Chaskey_a:=Chaskey_input_pi[2];   //<<< 16
   	Chaskey_Temp:=0;
   	//left shift Chaskey_b=16 bits
   	Chaskey_Temp.16:=Chaskey_a.0;
   	Chaskey_Temp.17:=Chaskey_a.1;
   	Chaskey_Temp.18:=Chaskey_a.2;
   	Chaskey_Temp.19:=Chaskey_a.3;
   	Chaskey_Temp.20:=Chaskey_a.4;
   	Chaskey_Temp.21:=Chaskey_a.5;
   	Chaskey_Temp.22:=Chaskey_a.6;
   	Chaskey_Temp.23:=Chaskey_a.7;
   	Chaskey_Temp.24:=Chaskey_a.8;
   	Chaskey_Temp.25:=Chaskey_a.9;
   	Chaskey_Temp.26:=Chaskey_a.10;
   	Chaskey_Temp.27:=Chaskey_a.11;
   	Chaskey_Temp.28:=Chaskey_a.12;
   	Chaskey_Temp.29:=Chaskey_a.13;
   	Chaskey_Temp.30:=Chaskey_a.14;
   	Chaskey_Temp.31:=Chaskey_a.15;
   	Chaskey_Temp.0:=Chaskey_a.16;
   	Chaskey_Temp.1:=Chaskey_a.17;
   	Chaskey_Temp.2:=Chaskey_a.18;
   	Chaskey_Temp.3:=Chaskey_a.19;
   	Chaskey_Temp.4:=Chaskey_a.20;
   	Chaskey_Temp.5:=Chaskey_a.21;
   	Chaskey_Temp.6:=Chaskey_a.22;
   	Chaskey_Temp.7:=Chaskey_a.23;
   	Chaskey_Temp.8:=Chaskey_a.24;
   	Chaskey_Temp.9:=Chaskey_a.25;
   	Chaskey_Temp.10:=Chaskey_a.26;
   	Chaskey_Temp.11:=Chaskey_a.27;
   	Chaskey_Temp.12:=Chaskey_a.28;
   	Chaskey_Temp.13:=Chaskey_a.29;
   	Chaskey_Temp.14:=Chaskey_a.30;
   	Chaskey_Temp.15:=Chaskey_a.31;
   	Chaskey_input_pi[2]:=Chaskey_Temp;
   end_for;
   
   
END_ROUTINE

ROUTINE If256   (* structured text *)
   	If OWF_Input[0].[0] Then
   		OWF_Result[0]:=OWF_Result[0] + 797041208+OWF_Add_c;
   		OWF_Add_c.0:=OWF_Result[0].31;
   		OWF_Result[0].31:=0;
   		OWF_Result[1]:=OWF_Result[1] + 1892147607+OWF_Add_c;
   		OWF_Add_c.1:=OWF_Result[1].31;
   		OWF_Result[1].31:=0;
   		OWF_Result[2]:=OWF_Result[2] + 272201627+OWF_Add_c;
   		OWF_Add_c.2:=OWF_Result[2].31;
   		OWF_Result[2].31:=0;
   		OWF_Result[3]:=OWF_Result[3] + 929594953+OWF_Add_c;
   		OWF_Add_c.3:=OWF_Result[3].31;
   		OWF_Result[3].31:=0;
   		OWF_Result[4]:=OWF_Result[4] + 1701098557+OWF_Add_c;
   		OWF_Add_c.4:=OWF_Result[4].31;
   		OWF_Result[4].31:=0;
   		OWF_Result[5]:=OWF_Result[5] + 1984918657+OWF_Add_c;
   		OWF_Add_c.5:=OWF_Result[5].31;
   		OWF_Result[5].31:=0;
   		OWF_Result[6]:=OWF_Result[6] + 2042310912+OWF_Add_c;
   		OWF_Add_c.6:=OWF_Result[6].31;
   		OWF_Result[6].31:=0;
   		OWF_Result[7]:=OWF_Result[7] + 1256180149+OWF_Add_c;
   		OWF_Add_c.7:=OWF_Result[7].31;
   		OWF_Result[7].31:=0;
   		OWF_Result[8]:=OWF_Result[8] + 2085759430+OWF_Add_c;
   		OWF_Add_c.8:=OWF_Result[8].31;
   		OWF_Result[8].31:=0;
   	End_If;
   	If OWF_Input[0].[1] Then
   		OWF_Result[0]:=OWF_Result[0] + 891262048+OWF_Add_c;
   		OWF_Add_c.0:=OWF_Result[0].31;
   		OWF_Result[0].31:=0;
   		OWF_Result[1]:=OWF_Result[1] + 1913322646+OWF_Add_c;
   		OWF_Add_c.1:=OWF_Result[1].31;
   		OWF_Result[1].31:=0;
   		OWF_Result[2]:=OWF_Result[2] + 157248836+OWF_Add_c;
   		OWF_Add_c.2:=OWF_Result[2].31;
   		OWF_Result[2].31:=0;
   		OWF_Result[3]:=OWF_Result[3] + 884867342+OWF_Add_c;
   		OWF_Add_c.3:=OWF_Result[3].31;
   		OWF_Result[3].31:=0;
   		OWF_Result[4]:=OWF_Result[4] + 188673317+OWF_Add_c;
   		OWF_Add_c.4:=OWF_Result[4].31;
   		OWF_Result[4].31:=0;
   		OWF_Result[5]:=OWF_Result[5] + 2096119266+OWF_Add_c;
   		OWF_Add_c.5:=OWF_Result[5].31;
   		OWF_Result[5].31:=0;
   		OWF_Result[6]:=OWF_Result[6] + 1480589067+OWF_Add_c;
   		OWF_Add_c.6:=OWF_Result[6].31;
   		OWF_Result[6].31:=0;
   		OWF_Result[7]:=OWF_Result[7] + 1099791289+OWF_Add_c;
   		OWF_Add_c.7:=OWF_Result[7].31;
   		OWF_Result[7].31:=0;
   		OWF_Result[8]:=OWF_Result[8] + 689702077+OWF_Add_c;
   		OWF_Add_c.8:=OWF_Result[8].31;
   		OWF_Result[8].31:=0;
   	End_If;
   	If OWF_Input[0].[2] Then
   		OWF_Result[0]:=OWF_Result[0] + 423846607+OWF_Add_c;
   		OWF_Add_c.0:=OWF_Result[0].31;
   		OWF_Result[0].31:=0;
   		OWF_Result[1]:=OWF_Result[1] + 221427001+OWF_Add_c;
   		OWF_Add_c.1:=OWF_Result[1].31;
   		OWF_Result[1].31:=0;
   		OWF_Result[2]:=OWF_Result[2] + 1557337489+OWF_Add_c;
   		OWF_Add_c.2:=OWF_Result[2].31;
   		OWF_Result[2].31:=0;
   		OWF_Result[3]:=OWF_Result[3] + 1284447123+OWF_Add_c;
   		OWF_Add_c.3:=OWF_Result[3].31;
   		OWF_Result[3].31:=0;
   		OWF_Result[4]:=OWF_Result[4] + 50932126+OWF_Add_c;
   		OWF_Add_c.4:=OWF_Result[4].31;
   		OWF_Result[4].31:=0;
   		OWF_Result[5]:=OWF_Result[5] + 49526266+OWF_Add_c;
   		OWF_Add_c.5:=OWF_Result[5].31;
   		OWF_Result[5].31:=0;
   		OWF_Result[6]:=OWF_Result[6] + 1509110851+OWF_Add_c;
   		OWF_Add_c.6:=OWF_Result[6].31;
   		OWF_Result[6].31:=0;
   		OWF_Result[7]:=OWF_Result[7] + 1330799634+OWF_Add_c;
   		OWF_Add_c.7:=OWF_Result[7].31;
   		OWF_Result[7].31:=0;
   		OWF_Result[8]:=OWF_Result[8] + 1410332622+OWF_Add_c;
   		OWF_Add_c.8:=OWF_Result[8].31;
   		OWF_Result[8].31:=0;
   	End_If;
   	If OWF_Input[0].[3] Then
   		OWF_Result[0]:=OWF_Result[0] + 1586608599+OWF_Add_c;
   		OWF_Add_c.0:=OWF_Result[0].31;
   		OWF_Result[0].31:=0;
   		OWF_Result[1]:=OWF_Result[1] + 1008757281+OWF_Add_c;
   		OWF_Add_c.1:=OWF_Result[1].31;
   		OWF_Result[1].31:=0;
   		OWF_Result[2]:=OWF_Result[2] + 1484532970+OWF_Add_c;
   		OWF_Add_c.2:=OWF_Result[2].31;
   		OWF_Result[2].31:=0;
   		OWF_Result[3]:=OWF_Result[3] + 793875947+OWF_Add_c;
   		OWF_Add_c.3:=OWF_Result[3].31;
   		OWF_Result[3].31:=0;
   		OWF_Result[4]:=OWF_Result[4] + 985404342+OWF_Add_c;
   		OWF_Add_c.4:=OWF_Result[4].31;
   		OWF_Result[4].31:=0;
   		OWF_Result[5]:=OWF_Result[5] + 1514352777+OWF_Add_c;
   		OWF_Add_c.5:=OWF_Result[5].31;
   		OWF_Result[5].31:=0;
   		OWF_Result[6]:=OWF_Result[6] + 1135345751+OWF_Add_c;
   		OWF_Add_c.6:=OWF_Result[6].31;
   		OWF_Result[6].31:=0;
   		OWF_Result[7]:=OWF_Result[7] + 672862598+OWF_Add_c;
   		OWF_Add_c.7:=OWF_Result[7].31;
   		OWF_Result[7].31:=0;
   		OWF_Result[8]:=OWF_Result[8] + 1484675889+OWF_Add_c;
   		OWF_Add_c.8:=OWF_Result[8].31;
   		OWF_Result[8].31:=0;
   	End_If;
   	If OWF_Input[0].[4] Then
   		OWF_Result[0]:=OWF_Result[0] + 614517358+OWF_Add_c;
   		OWF_Add_c.0:=OWF_Result[0].31;
   		OWF_Result[0].31:=0;
   		OWF_Result[1]:=OWF_Result[1] + 1070547517+OWF_Add_c;
   		OWF_Add_c.1:=OWF_Result[1].31;
   		OWF_Result[1].31:=0;
   		OWF_Result[2]:=OWF_Result[2] + 690174946+OWF_Add_c;
   		OWF_Add_c.2:=OWF_Result[2].31;
   		OWF_Result[2].31:=0;
   		OWF_Result[3]:=OWF_Result[3] + 889943012+OWF_Add_c;
   		OWF_Add_c.3:=OWF_Result[3].31;
   		OWF_Result[3].31:=0;
   		OWF_Result[4]:=OWF_Result[4] + 347648387+OWF_Add_c;
   		OWF_Add_c.4:=OWF_Result[4].31;
   		OWF_Result[4].31:=0;
   		OWF_Result[5]:=OWF_Result[5] + 1128332508+OWF_Add_c;
   		OWF_Add_c.5:=OWF_Result[5].31;
   		OWF_Result[5].31:=0;
   		OWF_Result[6]:=OWF_Result[6] + 1399662720+OWF_Add_c;
   		OWF_Add_c.6:=OWF_Result[6].31;
   		OWF_Result[6].31:=0;
   		OWF_Result[7]:=OWF_Result[7] + 1565377655+OWF_Add_c;
   		OWF_Add_c.7:=OWF_Result[7].31;
   		OWF_Result[7].31:=0;
   		OWF_Result[8]:=OWF_Result[8] + 1814409302+OWF_Add_c;
   		OWF_Add_c.8:=OWF_Result[8].31;
   		OWF_Result[8].31:=0;
   	End_If;
   	If OWF_Input[0].[5] Then
   		OWF_Result[0]:=OWF_Result[0] + 1800759771+OWF_Add_c;
   		OWF_Add_c.0:=OWF_Result[0].31;
   		OWF_Result[0].31:=0;
   		OWF_Result[1]:=OWF_Result[1] + 1223016147+OWF_Add_c;
   		OWF_Add_c.1:=OWF_Result[1].31;
   		OWF_Result[1].31:=0;
   		OWF_Result[2]:=OWF_Result[2] + 1501112628+OWF_Add_c;
   		OWF_Add_c.2:=OWF_Result[2].31;
   		OWF_Result[2].31:=0;
   		OWF_Result[3]:=OWF_Result[3] + 1971699393+OWF_Add_c;
   		OWF_Add_c.3:=OWF_Result[3].31;
   		OWF_Result[3].31:=0;
   		OWF_Result[4]:=OWF_Result[4] + 214300319+OWF_Add_c;
   		OWF_Add_c.4:=OWF_Result[4].31;
   		OWF_Result[4].31:=0;
   		OWF_Result[5]:=OWF_Result[5] + 1123701424+OWF_Add_c;
   		OWF_Add_c.5:=OWF_Result[5].31;
   		OWF_Result[5].31:=0;
   		OWF_Result[6]:=OWF_Result[6] + 155794511+OWF_Add_c;
   		OWF_Add_c.6:=OWF_Result[6].31;
   		OWF_Result[6].31:=0;
   		OWF_Result[7]:=OWF_Result[7] + 377658125+OWF_Add_c;
   		OWF_Add_c.7:=OWF_Result[7].31;
   		OWF_Result[7].31:=0;
   		OWF_Result[8]:=OWF_Result[8] + 1300678313+OWF_Add_c;
   		OWF_Add_c.8:=OWF_Result[8].31;
   		OWF_Result[8].31:=0;
   	End_If;
   	If OWF_Input[0].[6] Then
   		OWF_Result[0]:=OWF_Result[0] + 1247510715+OWF_Add_c;
   		OWF_Add_c.0:=OWF_Result[0].31;
   		OWF_Result[0].31:=0;
   		OWF_Result[1]:=OWF_Result[1] + 736041892+OWF_Add_c;
   		OWF_Add_c.1:=OWF_Result[1].31;
   		OWF_Result[1].31:=0;
   		OWF_Result[2]:=OWF_Result[2] + 898033892+OWF_Add_c;
   		OWF_Add_c.2:=OWF_Result[2].31;
   		OWF_Result[2].31:=0;
   		OWF_Result[3]:=OWF_Result[3] + 785690422+OWF_Add_c;
   		OWF_Add_c.3:=OWF_Result[3].31;
   		OWF_Result[3].31:=0;
   		OWF_Result[4]:=OWF_Result[4] + 309775084+OWF_Add_c;
   		OWF_Add_c.4:=OWF_Result[4].31;
   		OWF_Result[4].31:=0;
   		OWF_Result[5]:=OWF_Result[5] + 1644704994+OWF_Add_c;
   		OWF_Add_c.5:=OWF_Result[5].31;
   		OWF_Result[5].31:=0;
   		OWF_Result[6]:=OWF_Result[6] + 657852096+OWF_Add_c;
   		OWF_Add_c.6:=OWF_Result[6].31;
   		OWF_Result[6].31:=0;
   		OWF_Result[7]:=OWF_Result[7] + 469630175+OWF_Add_c;
   		OWF_Add_c.7:=OWF_Result[7].31;